REGION Network 5: Aggiorno mesaggio per richiesta di stato SCHEDA DELAY
   // ADDR+LRC
   RUNG wire#powerrail
      { S7_Templates := "SrcType := Word" } EQ_Contact(in1 := "SERIAL_DATA".ADDRESS, in2 := #INDIRIZZO_AQN)
      { S7_Templates := "SrcType := Word" } EQ_Contact(in1 := #comando_attivo, in2 := 0)
      Move(in := 16#00, out1 => "SERIAL_DATA".messaggio_76h[1])
      Move(in := 16#76, out1 => "SERIAL_DATA".messaggio_76h[4])
   END_RUNG
   // the same network as SCL:
   IF ("SERIAL_DATA".ADDRESS = #INDIRIZZO_AQN) AND (#comando_attivo = 0) THEN
       "SERIAL_DATA".messaggio_76h[1] := 16#00;
       "SERIAL_DATA".messaggio_76h[4] := 16#76;
   END_IF;
END_REGION

REGION Network 6: Aggiorno mesaggio per reset SCHEDA DELAY
   // ADDR+LRC
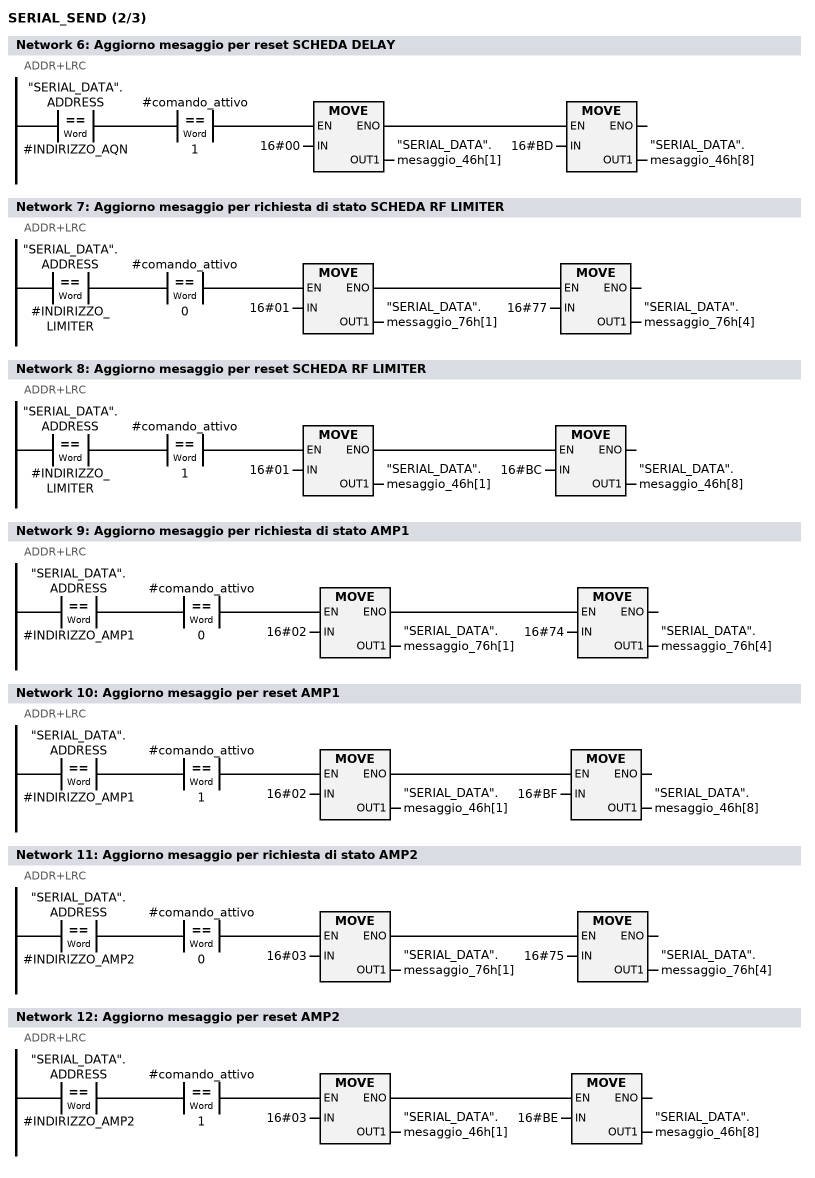
   RUNG wire#powerrail
      { S7_Templates := "SrcType := Word" } EQ_Contact(in1 := "SERIAL_DATA".ADDRESS, in2 := #INDIRIZZO_AQN)
      { S7_Templates := "SrcType := Word" } EQ_Contact(in1 := #comando_attivo, in2 := 1)
      Move(in := 16#00, out1 => "SERIAL_DATA".mesaggio_46h[1])
      Move(in := 16#BD, out1 => "SERIAL_DATA".mesaggio_46h[8])
   END_RUNG
   // the same network as SCL:
   IF ("SERIAL_DATA".ADDRESS = #INDIRIZZO_AQN) AND (#comando_attivo = 1) THEN
       "SERIAL_DATA".mesaggio_46h[1] := 16#00;
       "SERIAL_DATA".mesaggio_46h[8] := 16#BD;
   END_IF;
END_REGION

REGION Network 7: Aggiorno mesaggio per richiesta di stato SCHEDA RF LIMITER
   // ADDR+LRC
   RUNG wire#powerrail
      { S7_Templates := "SrcType := Word" } EQ_Contact(in1 := "SERIAL_DATA".ADDRESS, in2 := #INDIRIZZO_LIMITER)
      { S7_Templates := "SrcType := Word" } EQ_Contact(in1 := #comando_attivo, in2 := 0)
      Move(in := 16#01, out1 => "SERIAL_DATA".messaggio_76h[1])
      Move(in := 16#77, out1 => "SERIAL_DATA".messaggio_76h[4])
   END_RUNG
   // the same network as SCL:
   IF ("SERIAL_DATA".ADDRESS = #INDIRIZZO_LIMITER) AND (#comando_attivo = 0) THEN
       "SERIAL_DATA".messaggio_76h[1] := 16#01;
       "SERIAL_DATA".messaggio_76h[4] := 16#77;
   END_IF;
END_REGION

REGION Network 8: Aggiorno mesaggio per reset SCHEDA RF LIMITER
   // ADDR+LRC
   RUNG wire#powerrail
      { S7_Templates := "SrcType := Word" } EQ_Contact(in1 := "SERIAL_DATA".ADDRESS, in2 := #INDIRIZZO_LIMITER)
      { S7_Templates := "SrcType := Word" } EQ_Contact(in1 := #comando_attivo, in2 := 1)
      Move(in := 16#01, out1 => "SERIAL_DATA".mesaggio_46h[1])
      Move(in := 16#BC, out1 => "SERIAL_DATA".mesaggio_46h[8])
   END_RUNG
   // the same network as SCL:
   IF ("SERIAL_DATA".ADDRESS = #INDIRIZZO_LIMITER) AND (#comando_attivo = 1) THEN
       "SERIAL_DATA".mesaggio_46h[1] := 16#01;
       "SERIAL_DATA".mesaggio_46h[8] := 16#BC;
   END_IF;
END_REGION

REGION Network 9: Aggiorno mesaggio per richiesta di stato AMP1
   // ADDR+LRC
   RUNG wire#powerrail
      { S7_Templates := "SrcType := Word" } EQ_Contact(in1 := "SERIAL_DATA".ADDRESS, in2 := #INDIRIZZO_AMP1)
      { S7_Templates := "SrcType := Word" } EQ_Contact(in1 := #comando_attivo, in2 := 0)
      Move(in := 16#02, out1 => "SERIAL_DATA".messaggio_76h[1])
      Move(in := 16#74, out1 => "SERIAL_DATA".messaggio_76h[4])
   END_RUNG
   // the same network as SCL:
   IF ("SERIAL_DATA".ADDRESS = #INDIRIZZO_AMP1) AND (#comando_attivo = 0) THEN
       "SERIAL_DATA".messaggio_76h[1] := 16#02;
       "SERIAL_DATA".messaggio_76h[4] := 16#74;
   END_IF;
END_REGION

REGION Network 10: Aggiorno mesaggio per reset AMP1
   // ADDR+LRC
   RUNG wire#powerrail
      { S7_Templates := "SrcType := Word" } EQ_Contact(in1 := "SERIAL_DATA".ADDRESS, in2 := #INDIRIZZO_AMP1)
      { S7_Templates := "SrcType := Word" } EQ_Contact(in1 := #comando_attivo, in2 := 1)
      Move(in := 16#02, out1 => "SERIAL_DATA".mesaggio_46h[1])
      Move(in := 16#BF, out1 => "SERIAL_DATA".mesaggio_46h[8])
   END_RUNG
   // the same network as SCL:
   IF ("SERIAL_DATA".ADDRESS = #INDIRIZZO_AMP1) AND (#comando_attivo = 1) THEN
       "SERIAL_DATA".mesaggio_46h[1] := 16#02;
       "SERIAL_DATA".mesaggio_46h[8] := 16#BF;
   END_IF;
END_REGION

REGION Network 11: Aggiorno mesaggio per richiesta di stato AMP2
   // ADDR+LRC
   RUNG wire#powerrail
      { S7_Templates := "SrcType := Word" } EQ_Contact(in1 := "SERIAL_DATA".ADDRESS, in2 := #INDIRIZZO_AMP2)
      { S7_Templates := "SrcType := Word" } EQ_Contact(in1 := #comando_attivo, in2 := 0)
      Move(in := 16#03, out1 => "SERIAL_DATA".messaggio_76h[1])
      Move(in := 16#75, out1 => "SERIAL_DATA".messaggio_76h[4])
   END_RUNG
   // the same network as SCL:
   IF ("SERIAL_DATA".ADDRESS = #INDIRIZZO_AMP2) AND (#comando_attivo = 0) THEN
       "SERIAL_DATA".messaggio_76h[1] := 16#03;
       "SERIAL_DATA".messaggio_76h[4] := 16#75;
   END_IF;
END_REGION

REGION Network 12: Aggiorno mesaggio per reset AMP2
   // ADDR+LRC
   RUNG wire#powerrail
      { S7_Templates := "SrcType := Word" } EQ_Contact(in1 := "SERIAL_DATA".ADDRESS, in2 := #INDIRIZZO_AMP2)
      { S7_Templates := "SrcType := Word" } EQ_Contact(in1 := #comando_attivo, in2 := 1)
      Move(in := 16#03, out1 => "SERIAL_DATA".mesaggio_46h[1])
      Move(in := 16#BE, out1 => "SERIAL_DATA".mesaggio_46h[8])
   END_RUNG
   // the same network as SCL:
   IF ("SERIAL_DATA".ADDRESS = #INDIRIZZO_AMP2) AND (#comando_attivo = 1) THEN
       "SERIAL_DATA".mesaggio_46h[1] := 16#03;
       "SERIAL_DATA".mesaggio_46h[8] := 16#BE;
   END_IF;
END_REGION

REGION Network 13: Aggiorno mesaggio per richiesta di stato DRV
   // ADDR+LRC
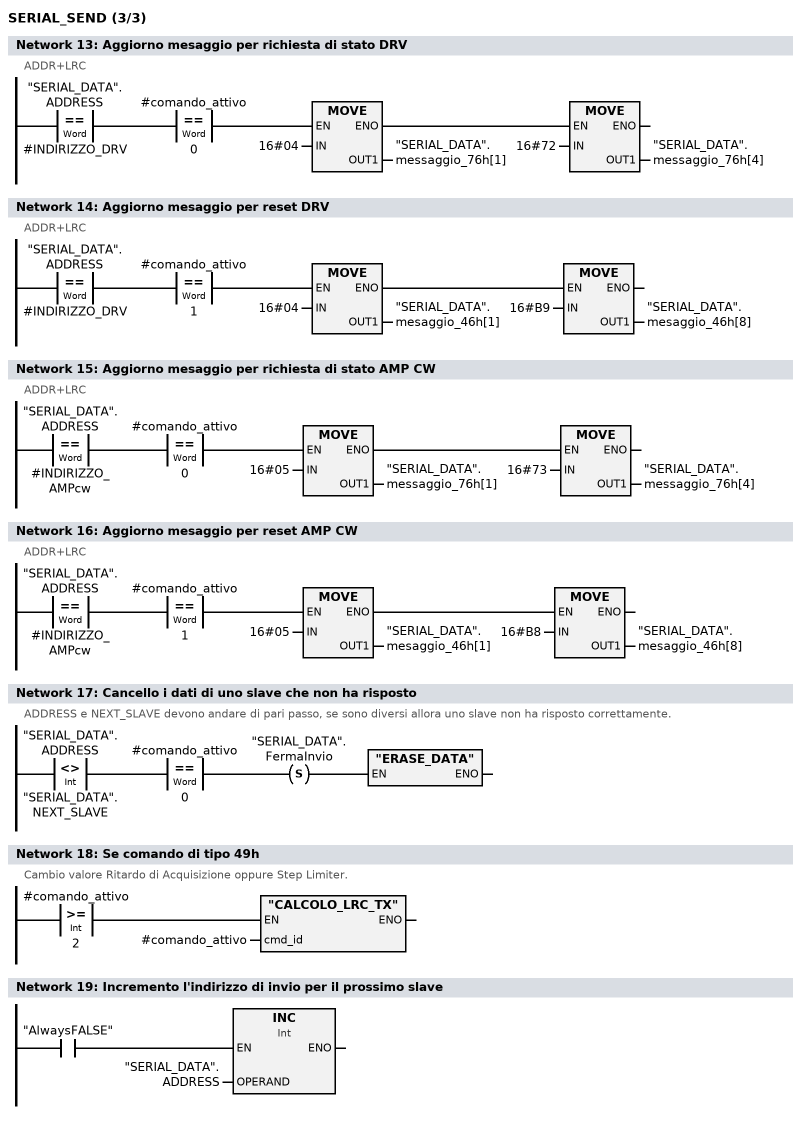
   RUNG wire#powerrail
      { S7_Templates := "SrcType := Word" } EQ_Contact(in1 := "SERIAL_DATA".ADDRESS, in2 := #INDIRIZZO_DRV)
      { S7_Templates := "SrcType := Word" } EQ_Contact(in1 := #comando_attivo, in2 := 0)
      Move(in := 16#04, out1 => "SERIAL_DATA".messaggio_76h[1])
      Move(in := 16#72, out1 => "SERIAL_DATA".messaggio_76h[4])
   END_RUNG
   // the same network as SCL:
   IF ("SERIAL_DATA".ADDRESS = #INDIRIZZO_DRV) AND (#comando_attivo = 0) THEN
       "SERIAL_DATA".messaggio_76h[1] := 16#04;
       "SERIAL_DATA".messaggio_76h[4] := 16#72;
   END_IF;
END_REGION

REGION Network 14: Aggiorno mesaggio per reset DRV
   // ADDR+LRC
   RUNG wire#powerrail
      { S7_Templates := "SrcType := Word" } EQ_Contact(in1 := "SERIAL_DATA".ADDRESS, in2 := #INDIRIZZO_DRV)
      { S7_Templates := "SrcType := Word" } EQ_Contact(in1 := #comando_attivo, in2 := 1)
      Move(in := 16#04, out1 => "SERIAL_DATA".mesaggio_46h[1])
      Move(in := 16#B9, out1 => "SERIAL_DATA".mesaggio_46h[8])
   END_RUNG
   // the same network as SCL:
   IF ("SERIAL_DATA".ADDRESS = #INDIRIZZO_DRV) AND (#comando_attivo = 1) THEN
       "SERIAL_DATA".mesaggio_46h[1] := 16#04;
       "SERIAL_DATA".mesaggio_46h[8] := 16#B9;
   END_IF;
END_REGION

REGION Network 15: Aggiorno mesaggio per richiesta di stato AMP CW
   // ADDR+LRC
   RUNG wire#powerrail
      { S7_Templates := "SrcType := Word" } EQ_Contact(in1 := "SERIAL_DATA".ADDRESS, in2 := #INDIRIZZO_AMPcw)
      { S7_Templates := "SrcType := Word" } EQ_Contact(in1 := #comando_attivo, in2 := 0)
      Move(in := 16#05, out1 => "SERIAL_DATA".messaggio_76h[1])
      Move(in := 16#73, out1 => "SERIAL_DATA".messaggio_76h[4])
   END_RUNG
   // the same network as SCL:
   IF ("SERIAL_DATA".ADDRESS = #INDIRIZZO_AMPcw) AND (#comando_attivo = 0) THEN
       "SERIAL_DATA".messaggio_76h[1] := 16#05;
       "SERIAL_DATA".messaggio_76h[4] := 16#73;
   END_IF;
END_REGION

REGION Network 16: Aggiorno mesaggio per reset AMP CW
   // ADDR+LRC
   RUNG wire#powerrail
      { S7_Templates := "SrcType := Word" } EQ_Contact(in1 := "SERIAL_DATA".ADDRESS, in2 := #INDIRIZZO_AMPcw)
      { S7_Templates := "SrcType := Word" } EQ_Contact(in1 := #comando_attivo, in2 := 1)
      Move(in := 16#05, out1 => "SERIAL_DATA".mesaggio_46h[1])
      Move(in := 16#B8, out1 => "SERIAL_DATA".mesaggio_46h[8])
   END_RUNG
   // the same network as SCL:
   IF ("SERIAL_DATA".ADDRESS = #INDIRIZZO_AMPcw) AND (#comando_attivo = 1) THEN
       "SERIAL_DATA".mesaggio_46h[1] := 16#05;
       "SERIAL_DATA".mesaggio_46h[8] := 16#B8;
   END_IF;
END_REGION

REGION Network 17: Cancello i dati di uno slave che non ha risposto
   // ADDRESS e NEXT_SLAVE devono andare di pari passo, se sono diversi allora uno slave non ha risposto correttamente.
   RUNG wire#powerrail
      { S7_Templates := "SrcType := Int" } NE_Contact(in1 := "SERIAL_DATA".ADDRESS, in2 := "SERIAL_DATA".NEXT_SLAVE)
      { S7_Templates := "SrcType := Word" } EQ_Contact(in1 := #comando_attivo, in2 := 0)
      S_Coil( "SERIAL_DATA".FermaInvio )
      "ERASE_DATA"()
   END_RUNG
   // the same network as SCL:
   IF ("SERIAL_DATA".ADDRESS <> "SERIAL_DATA".NEXT_SLAVE) AND (#comando_attivo = 0) THEN
       "SERIAL_DATA".FermaInvio := TRUE;
       "ERASE_DATA"();
   END_IF;
END_REGION

REGION Network 18: Se comando di tipo 49h
   // Cambio valore Ritardo di Acquisizione oppure Step Limiter.
   RUNG wire#powerrail
      { S7_Templates := "SrcType := Int" } GE_Contact(in1 := #comando_attivo, in2 := 2)
      "CALCOLO_LRC_TX"(cmd_id := #comando_attivo)
   END_RUNG
   // the same network as SCL:
   IF #comando_attivo >= 2 THEN "CALCOLO_LRC_TX"(cmd_id := #comando_attivo); END_IF;
END_REGION

REGION Network 19: Incremento l'indirizzo di invio per il prossimo slave
   RUNG wire#powerrail
      Contact( "AlwaysFALSE" )
      { S7_Templates := "DestType := Int" } Inc( "SERIAL_DATA".ADDRESS )
   END_RUNG
   // the same network as SCL:
   IF "AlwaysFALSE" THEN "SERIAL_DATA".ADDRESS := "SERIAL_DATA".ADDRESS + 1; END_IF;
END_REGION
END_FUNCTION

FUNCTION "SERIAL_RECEIVE" : Void   // FC4, LAD
TITLE = SERIAL RECEIVE
{ S7_Optimized_Access := 'FALSE' }
VERSION : 0.1
   VAR_TEMP   // added for the SCL form of the ladder/FBD networks
      _w1 : Bool;
   END_VAR
BEGIN

REGION Network 1: Calcolo LRC del messaggio ricevuto
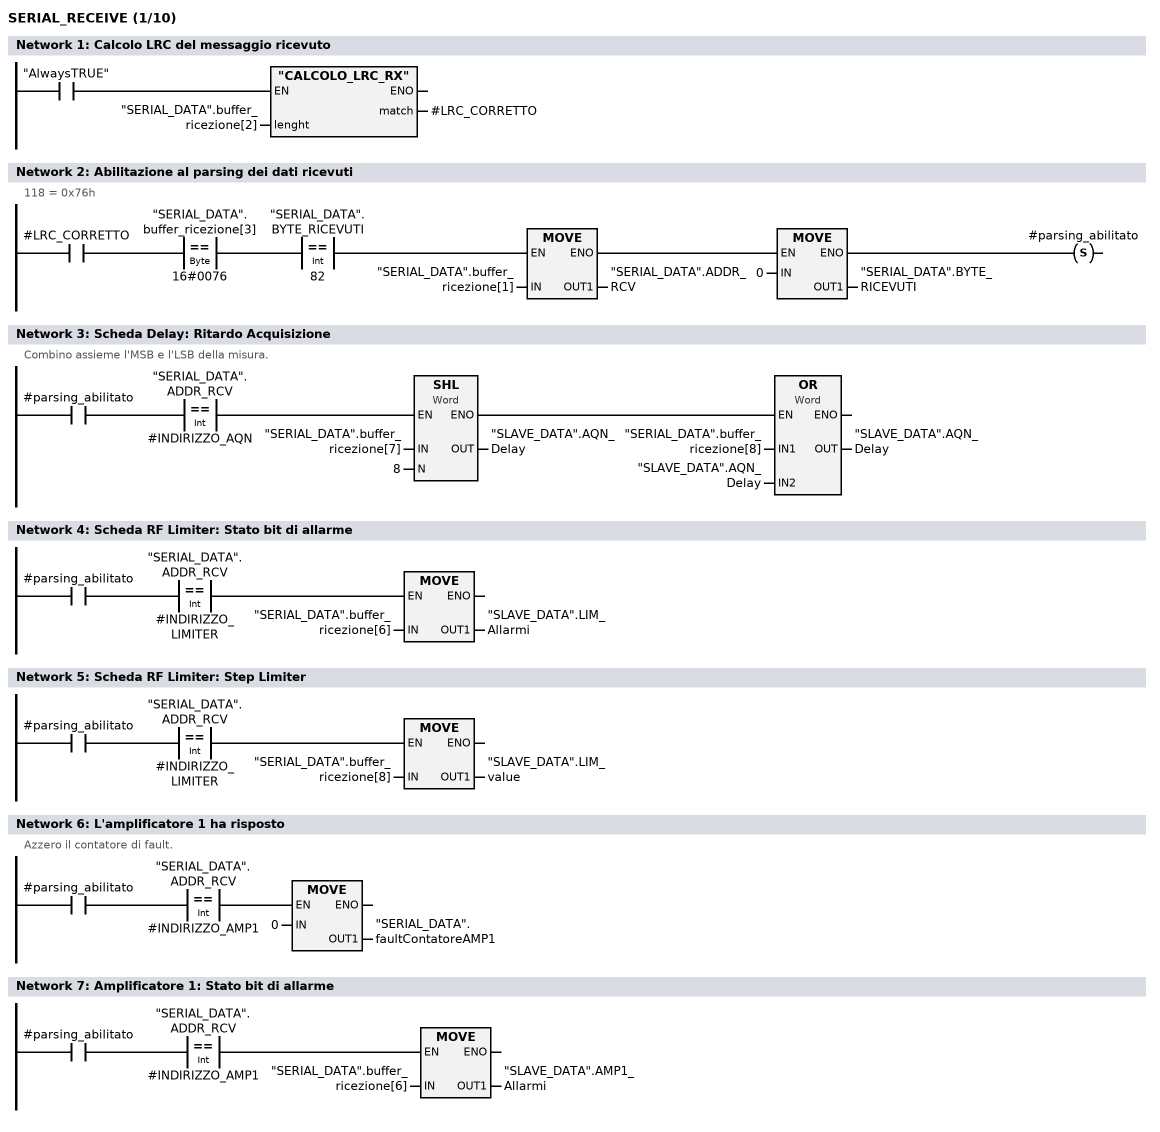
   RUNG wire#powerrail
      Contact( "AlwaysTRUE" )
      "CALCOLO_LRC_RX"(lenght := "SERIAL_DATA".buffer_ricezione[2], match => #LRC_CORRETTO)
   END_RUNG
   // the same network as SCL:
   IF "AlwaysTRUE" THEN
       "CALCOLO_LRC_RX"(lenght := "SERIAL_DATA".buffer_ricezione[2], match => #LRC_CORRETTO);
   END_IF;
END_REGION

REGION Network 2: Abilitazione al parsing dei dati ricevuti
   // 118 = 0x76h
   RUNG wire#powerrail
      Contact( #LRC_CORRETTO )
      { S7_Templates := "SrcType := Byte" } EQ_Contact(in1 := "SERIAL_DATA".buffer_ricezione[3], in2 := 16#0076)
      { S7_Templates := "SrcType := Int" } EQ_Contact(in1 := "SERIAL_DATA".BYTE_RICEVUTI, in2 := 82)
      Move(in := "SERIAL_DATA".buffer_ricezione[1], out1 => "SERIAL_DATA".ADDR_RCV)
      Move(in := 0, out1 => "SERIAL_DATA".BYTE_RICEVUTI)
      S_Coil( #parsing_abilitato )
   END_RUNG
   // the same network as SCL:
   IF #LRC_CORRETTO AND ("SERIAL_DATA".buffer_ricezione[3] = 16#0076) AND ("SERIAL_DATA".BYTE_RICEVUTI = 82) THEN
       "SERIAL_DATA".ADDR_RCV := "SERIAL_DATA".buffer_ricezione[1];
   END_IF;
   #_w1 := #LRC_CORRETTO AND ("SERIAL_DATA".buffer_ricezione[3] = 16#0076) AND ("SERIAL_DATA".BYTE_RICEVUTI = 82);
   IF #_w1 THEN
       "SERIAL_DATA".BYTE_RICEVUTI := 0;
       #parsing_abilitato := TRUE;
   END_IF;
END_REGION

REGION Network 3: Scheda Delay: Ritardo Acquisizione
   // Combino assieme l'MSB e l'LSB della misura.
   // no checked SCL form for this network; see the picture
END_REGION

REGION Network 4: Scheda RF Limiter: Stato bit di allarme
   RUNG wire#powerrail
      Contact( #parsing_abilitato )
      { S7_Templates := "SrcType := Int" } EQ_Contact(in1 := "SERIAL_DATA".ADDR_RCV, in2 := #INDIRIZZO_LIMITER)
      Move(in := "SERIAL_DATA".buffer_ricezione[6], out1 => "SLAVE_DATA".LIM_Allarmi)
   END_RUNG
   // the same network as SCL:
   IF #parsing_abilitato AND ("SERIAL_DATA".ADDR_RCV = #INDIRIZZO_LIMITER) THEN
       "SLAVE_DATA".LIM_Allarmi := "SERIAL_DATA".buffer_ricezione[6];
   END_IF;
END_REGION

REGION Network 5: Scheda RF Limiter: Step Limiter
   RUNG wire#powerrail
      Contact( #parsing_abilitato )
      { S7_Templates := "SrcType := Int" } EQ_Contact(in1 := "SERIAL_DATA".ADDR_RCV, in2 := #INDIRIZZO_LIMITER)
      Move(in := "SERIAL_DATA".buffer_ricezione[8], out1 => "SLAVE_DATA".LIM_value)
   END_RUNG
   // the same network as SCL:
   IF #parsing_abilitato AND ("SERIAL_DATA".ADDR_RCV = #INDIRIZZO_LIMITER) THEN
       "SLAVE_DATA".LIM_value := "SERIAL_DATA".buffer_ricezione[8];
   END_IF;
END_REGION

REGION Network 6: L'amplificatore 1 ha risposto
   // Azzero il contatore di fault.
   RUNG wire#powerrail
      Contact( #parsing_abilitato )
      { S7_Templates := "SrcType := Int" } EQ_Contact(in1 := "SERIAL_DATA".ADDR_RCV, in2 := #INDIRIZZO_AMP1)
      Move(in := 0, out1 => "SERIAL_DATA".faultContatoreAMP1)
   END_RUNG
   // the same network as SCL:
   IF #parsing_abilitato AND ("SERIAL_DATA".ADDR_RCV = #INDIRIZZO_AMP1) THEN
       "SERIAL_DATA".faultContatoreAMP1 := 0;
   END_IF;
END_REGION

REGION Network 7: Amplificatore 1: Stato bit di allarme
   RUNG wire#powerrail
      Contact( #parsing_abilitato )
      { S7_Templates := "SrcType := Int" } EQ_Contact(in1 := "SERIAL_DATA".ADDR_RCV, in2 := #INDIRIZZO_AMP1)
      Move(in := "SERIAL_DATA".buffer_ricezione[6], out1 => "SLAVE_DATA".AMP1_Allarmi)
   END_RUNG
   // the same network as SCL:
   IF #parsing_abilitato AND ("SERIAL_DATA".ADDR_RCV = #INDIRIZZO_AMP1) THEN
       "SLAVE_DATA".AMP1_Allarmi := "SERIAL_DATA".buffer_ricezione[6];
   END_IF;
END_REGION

REGION Network 8: Amplificatore 1: V1
   // Combino assieme l'MSB e l'LSB della misura.
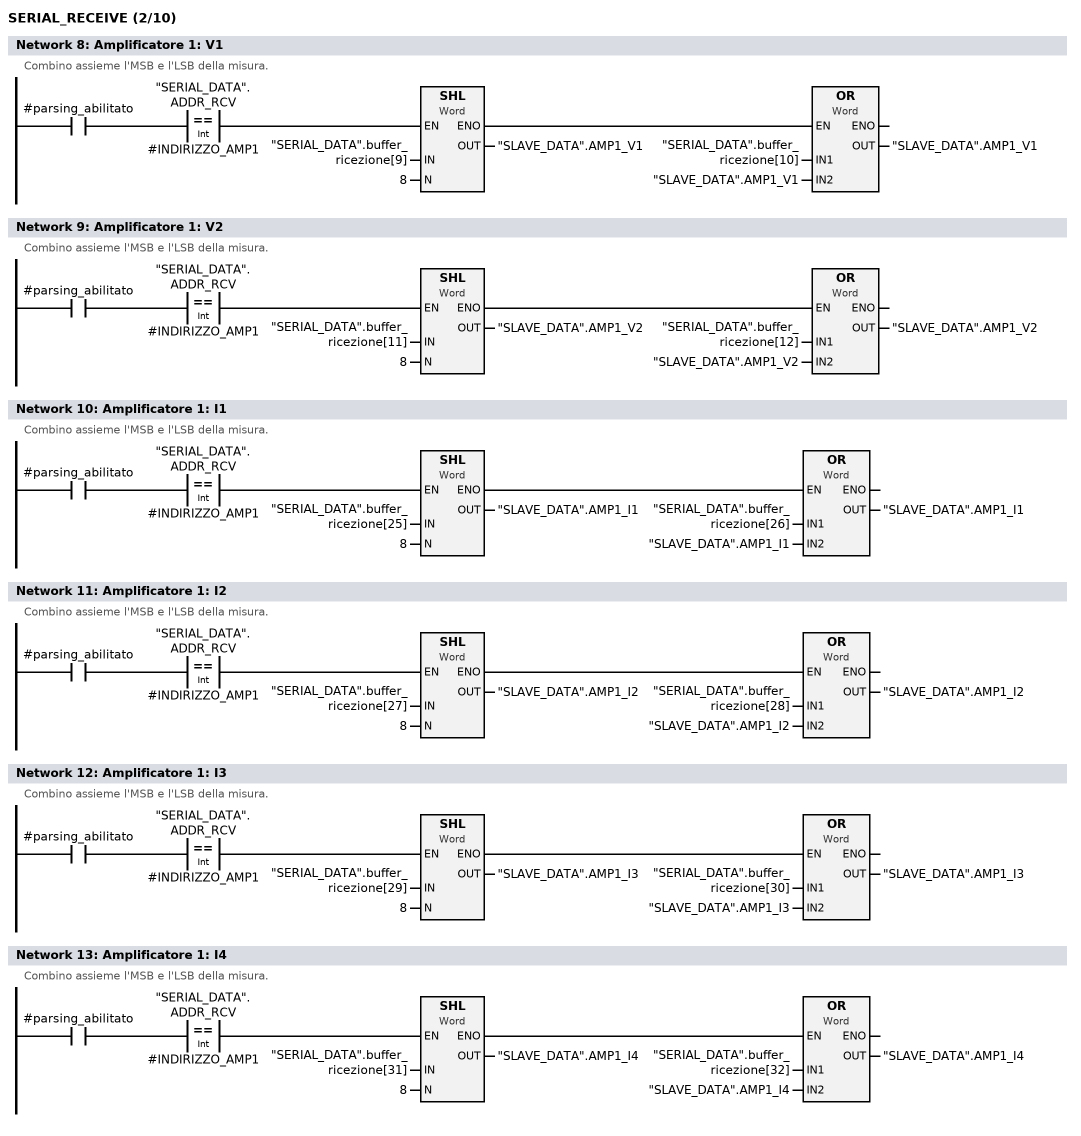
   // no checked SCL form for this network; see the picture
END_REGION

REGION Network 9: Amplificatore 1: V2
   // Combino assieme l'MSB e l'LSB della misura.
   // no checked SCL form for this network; see the picture
END_REGION

REGION Network 10: Amplificatore 1: I1
   // Combino assieme l'MSB e l'LSB della misura.
   // no checked SCL form for this network; see the picture
END_REGION

REGION Network 11: Amplificatore 1: I2
   // Combino assieme l'MSB e l'LSB della misura.
   // no checked SCL form for this network; see the picture
END_REGION

REGION Network 12: Amplificatore 1: I3
   // Combino assieme l'MSB e l'LSB della misura.
   // no checked SCL form for this network; see the picture
END_REGION

REGION Network 13: Amplificatore 1: I4
   // Combino assieme l'MSB e l'LSB della misura.
   // no checked SCL form for this network; see the picture
END_REGION

REGION Network 14: Amplificatore 1: I5
   // Combino assieme l'MSB e l'LSB della misura.
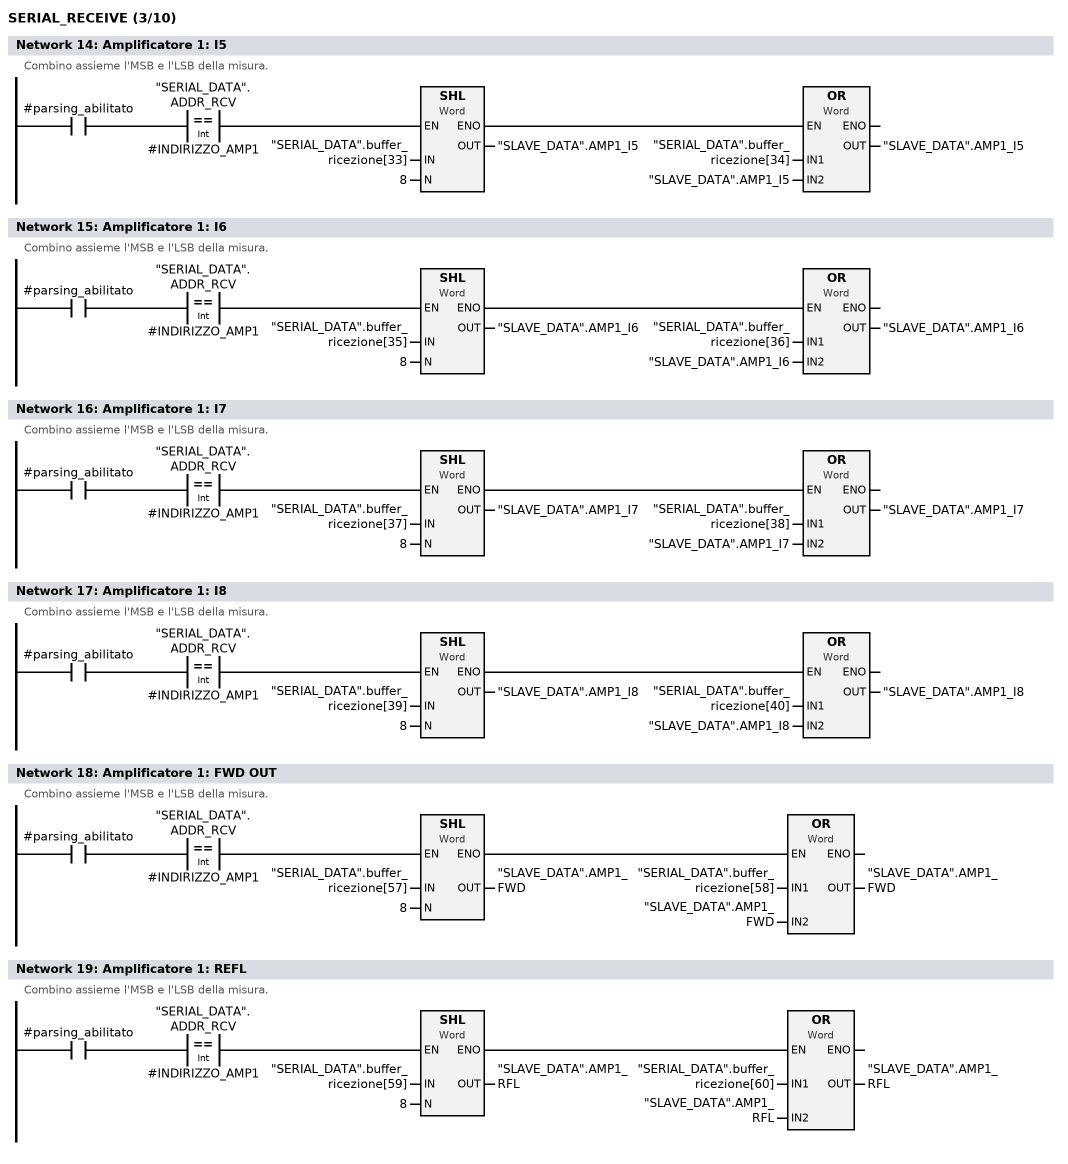
   // no checked SCL form for this network; see the picture
END_REGION

REGION Network 15: Amplificatore 1: I6
   // Combino assieme l'MSB e l'LSB della misura.
   // no checked SCL form for this network; see the picture
END_REGION

REGION Network 16: Amplificatore 1: I7
   // Combino assieme l'MSB e l'LSB della misura.
   // no checked SCL form for this network; see the picture
END_REGION

REGION Network 17: Amplificatore 1: I8
   // Combino assieme l'MSB e l'LSB della misura.
   // no checked SCL form for this network; see the picture
END_REGION

REGION Network 18: Amplificatore 1: FWD OUT
   // Combino assieme l'MSB e l'LSB della misura.
   // no checked SCL form for this network; see the picture
END_REGION

REGION Network 19: Amplificatore 1: REFL
   // Combino assieme l'MSB e l'LSB della misura.
   // no checked SCL form for this network; see the picture
END_REGION

REGION Network 20: Amplificatore 1: FWD IN
   // Combino assieme l'MSB e l'LSB della misura.
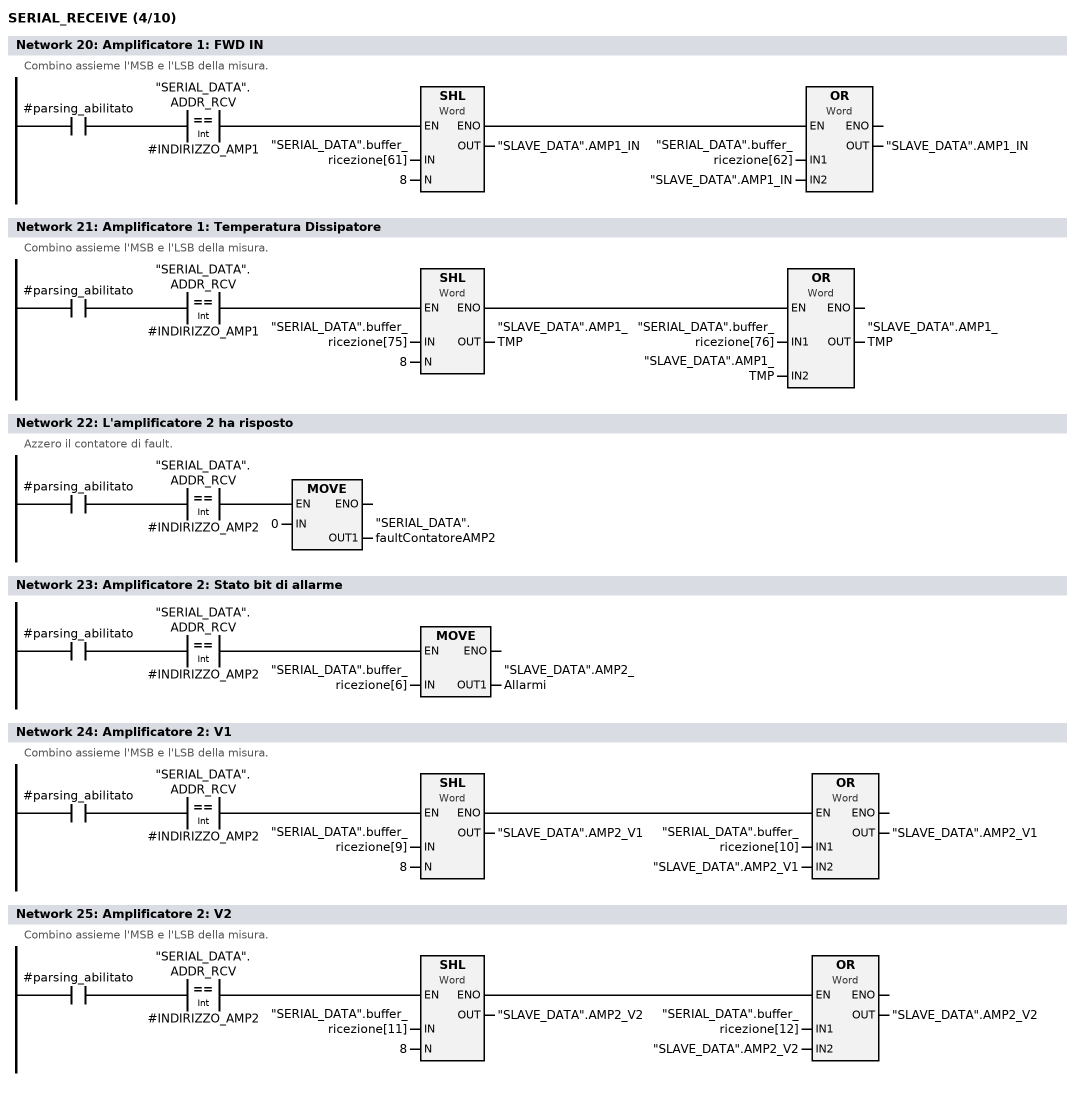
   // no checked SCL form for this network; see the picture
END_REGION

REGION Network 21: Amplificatore 1: Temperatura Dissipatore
   // Combino assieme l'MSB e l'LSB della misura.
   // no checked SCL form for this network; see the picture
END_REGION

REGION Network 22: L'amplificatore 2 ha risposto
   // Azzero il contatore di fault.
   RUNG wire#powerrail
      Contact( #parsing_abilitato )
      { S7_Templates := "SrcType := Int" } EQ_Contact(in1 := "SERIAL_DATA".ADDR_RCV, in2 := #INDIRIZZO_AMP2)
      Move(in := 0, out1 => "SERIAL_DATA".faultContatoreAMP2)
   END_RUNG
   // the same network as SCL:
   IF #parsing_abilitato AND ("SERIAL_DATA".ADDR_RCV = #INDIRIZZO_AMP2) THEN
       "SERIAL_DATA".faultContatoreAMP2 := 0;
   END_IF;
END_REGION

REGION Network 23: Amplificatore 2: Stato bit di allarme
   RUNG wire#powerrail
      Contact( #parsing_abilitato )
      { S7_Templates := "SrcType := Int" } EQ_Contact(in1 := "SERIAL_DATA".ADDR_RCV, in2 := #INDIRIZZO_AMP2)
      Move(in := "SERIAL_DATA".buffer_ricezione[6], out1 => "SLAVE_DATA".AMP2_Allarmi)
   END_RUNG
   // the same network as SCL:
   IF #parsing_abilitato AND ("SERIAL_DATA".ADDR_RCV = #INDIRIZZO_AMP2) THEN
       "SLAVE_DATA".AMP2_Allarmi := "SERIAL_DATA".buffer_ricezione[6];
   END_IF;
END_REGION

REGION Network 24: Amplificatore 2: V1
   // Combino assieme l'MSB e l'LSB della misura.
   // no checked SCL form for this network; see the picture
END_REGION

REGION Network 25: Amplificatore 2: V2
   // Combino assieme l'MSB e l'LSB della misura.
   // no checked SCL form for this network; see the picture
END_REGION

REGION Network 26: Amplificatore 2: I1
   // Combino assieme l'MSB e l'LSB della misura.
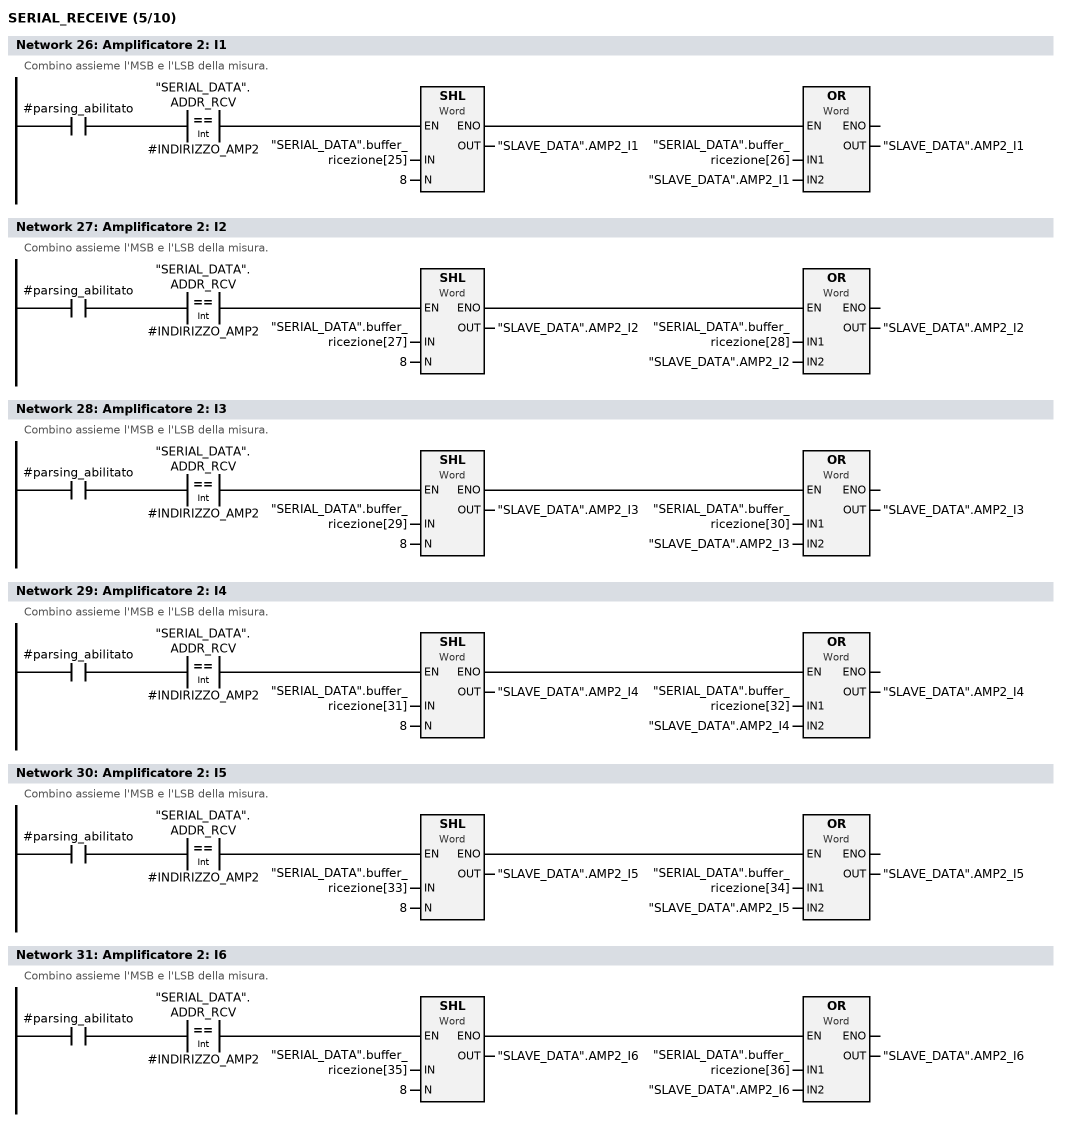
   // no checked SCL form for this network; see the picture
END_REGION

REGION Network 27: Amplificatore 2: I2
   // Combino assieme l'MSB e l'LSB della misura.
   // no checked SCL form for this network; see the picture
END_REGION

REGION Network 28: Amplificatore 2: I3
   // Combino assieme l'MSB e l'LSB della misura.
   // no checked SCL form for this network; see the picture
END_REGION

REGION Network 29: Amplificatore 2: I4
   // Combino assieme l'MSB e l'LSB della misura.
   // no checked SCL form for this network; see the picture
END_REGION

REGION Network 30: Amplificatore 2: I5
   // Combino assieme l'MSB e l'LSB della misura.
   // no checked SCL form for this network; see the picture
END_REGION

REGION Network 31: Amplificatore 2: I6
   // Combino assieme l'MSB e l'LSB della misura.
   // no checked SCL form for this network; see the picture
END_REGION

REGION Network 32: Amplificatore 2: I7
   // Combino assieme l'MSB e l'LSB della misura.
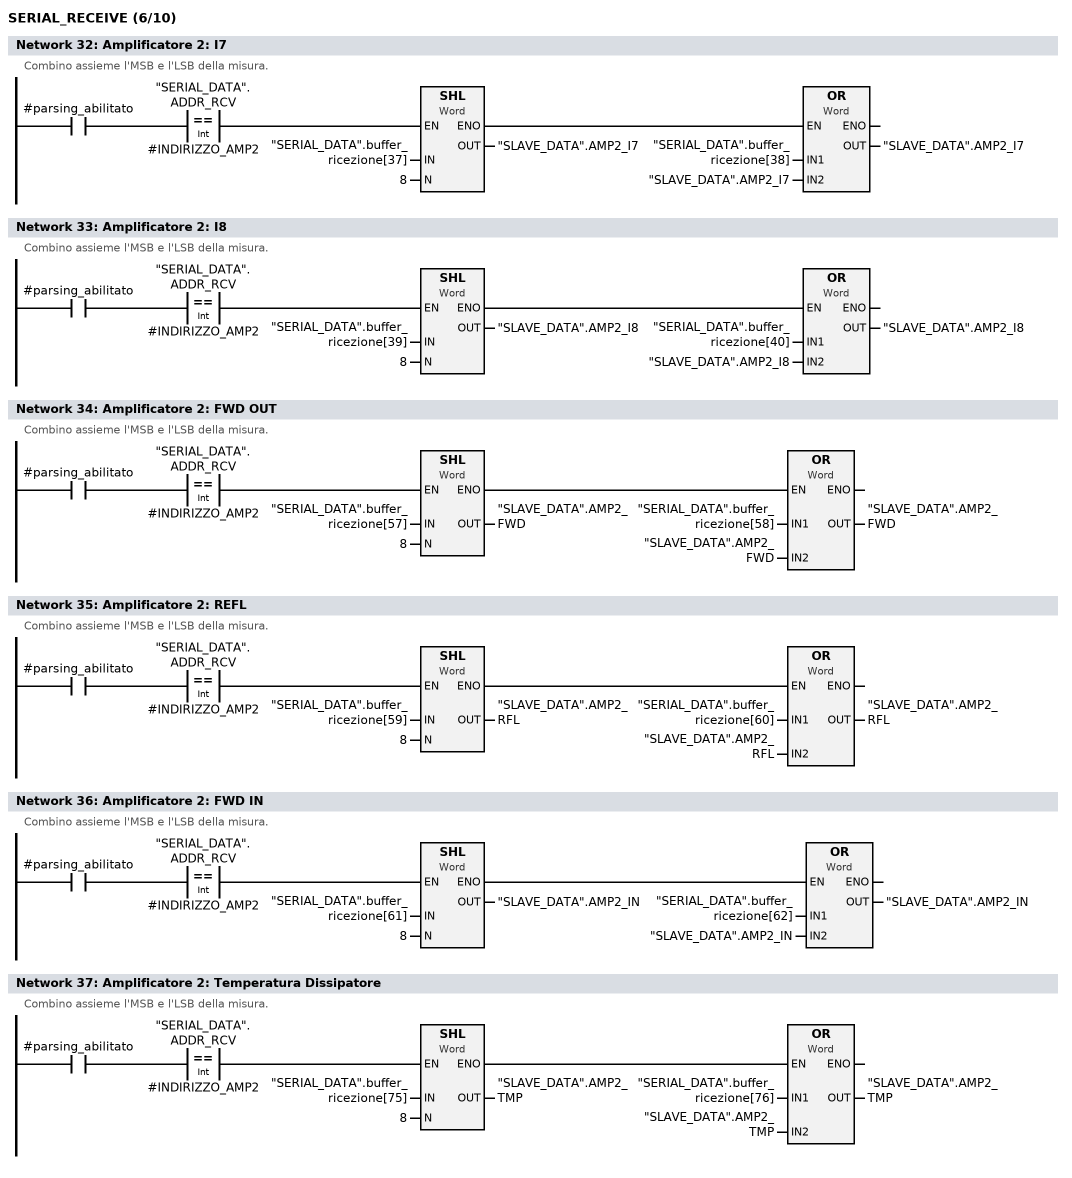
   // no checked SCL form for this network; see the picture
END_REGION

REGION Network 33: Amplificatore 2: I8
   // Combino assieme l'MSB e l'LSB della misura.
   // no checked SCL form for this network; see the picture
END_REGION

REGION Network 34: Amplificatore 2: FWD OUT
   // Combino assieme l'MSB e l'LSB della misura.
   // no checked SCL form for this network; see the picture
END_REGION

REGION Network 35: Amplificatore 2: REFL
   // Combino assieme l'MSB e l'LSB della misura.
   // no checked SCL form for this network; see the picture
END_REGION

REGION Network 36: Amplificatore 2: FWD IN
   // Combino assieme l'MSB e l'LSB della misura.
   // no checked SCL form for this network; see the picture
END_REGION

REGION Network 37: Amplificatore 2: Temperatura Dissipatore
   // Combino assieme l'MSB e l'LSB della misura.
   // no checked SCL form for this network; see the picture
END_REGION

REGION Network 38: Il driver ha risposto
   // Azzero il contatore di fault.